// TIA Portal project "inzynierka2" (V17)

(* hardware
DEVICE "S7-1500/ET200MP station_1"  S7-1500 station
   slot 0: "Rail_0"  Rack  6ES7 590-1***0-0AA0
   slot 1: "PLC_1"  CPU 1513-1 PN  6ES7 513-1AL00-0AB0  V1.1
      slot 3: "CPU display_1"  6ES7591-1XA00-0AA0
      slot 32768: "PROFINET interface_1"  X1
DEVICE "GSD device_1"  GSD.Device.PN
   slot 0: "Rack"  Rack  V1.0
   slot 0: "CPX"  CPX-RC  TN 197330  V3.2.24
      slot 0: "CPX-RC"  CPX-RC
      slot 1: "PN-IO Interface"  PN-IO Interface
         slot 1: "Port 1"  Port 1
         slot 2: "Port 2"  Port 2
   slot 1: "FB34 PNIO Module (RC) [8IB/8OB]_1"  FB34 PNIO Module (RC) [8IB/8OB]  TN 548751, CPX-FB34
      slot 0: "FB34 PNIO Module (RC) [8IB/8OB]"  FB34 PNIO Module (RC) [8IB/8OB]
DEVICE "HMI_1"  KTP700 Basic PN
   slot 0: "HMI_1"  KTP700 Basic PN  6AV2 123-2GB03-0AX0  15.0.0.0
   slot 1: "HMI_RT_1"  KTP700 Basic PN  6AV2 123-2GB03-0AX0  15.0.0.0
   slot 5: "HMI_1.IE_CP_1"  PROFINET Interface  15.0.0.0
      slot 1: "PROFINET Interface_1"  PROFINET Interface
         slot 1: "Port_1"  Port
*)

// ===== PLC "PLC_1"  CPU 1513-1 PN =====

VAR_GLOBAL   // PLC tag table "Default tag table"
   "System_Byte" AT %MB1 : Byte;
   "FirstScan" AT %M1.0 : Bool;
   "DiagStatusUpdate" AT %M1.1 : Bool;
   "AlwaysTRUE" AT %M1.2 : Bool;
   "AlwaysFALSE" AT %M1.3 : Bool;
   "Clock_Byte" AT %MB0 : Byte;
   "Clock_10Hz" AT %M0.0 : Bool;
   "Clock_5Hz" AT %M0.1 : Bool;
   "Clock_2.5Hz" AT %M0.2 : Bool;
   "Clock_2Hz" AT %M0.3 : Bool;
   "Clock_1.25Hz" AT %M0.4 : Bool;
   "Clock_1Hz" AT %M0.5 : Bool;
   "Clock_0.625Hz" AT %M0.6 : Bool;
   "Clock_0.5Hz" AT %M0.7 : Bool;
   "Tag_1" AT %M10.1 : Bool;
   "testowy" AT %MB20 : Byte;
   "testowy_out" AT %MB22 : Byte;
   "testowy2" AT %MB21 : Byte;
   "testowy_out2" AT %MB23 : Byte;
   "Tag_2" AT %IW0 : Word;
   "IB_MANOMETER1_2" AT %IB0 : Byte;
   "IB_MANOMETER1_1" AT %IB1 : Byte;
   "valves_out_1" AT %MB100 : Byte;
   "QB0_BYTE_OUT" AT %QB0 : Byte;
   "valves_out_2" AT %MB101 : Byte;
   "QB1_BYTE_OUT" AT %QB1 : Byte;
   "QB2_BYTE_VALVE_OPEN_TO_SEND" AT %QB2 : Byte;
   "IB_MANOMETER3_2" AT %IB2 : Byte;
   "IB_MANOMETER3_1" AT %IB3 : Byte;
   "testint" AT %MW210 : Int;
   "testhmibool" AT %M212.0 : Bool;
   "IB_VALVE_STATE_1" AT %IB4 : Byte;
   "IB_VALVE_STATE_2" AT %IB5 : Byte;
   "IB_VALVE_STATE_3" AT %IB6 : Byte;
   "IB_VALVE_STATE_4" AT %IB7 : Byte;
   "Tag_3" AT %IB8 : Byte;
END_VAR

DATA_BLOCK "DB_send_rcv"   // DB1
{ S7_Optimized_Access := 'TRUE' }
VERSION : 0.1
   VAR
      przesuniecie : USInt;
      BAJT1 : Byte;
      BAJT2 : Byte;
      MANOMETER1_VALUE : Real;
      MANOMETER3_VALUE : Real;
      VALVE_OPEN_PERCENT : Int;
   END_VAR
BEGIN
END_DATA_BLOCK

DATA_BLOCK "DB_valves"   // DB2
{ S7_Optimized_Access := 'TRUE' }
VERSION : 0.1
   VAR
      VALVEMODE : Int := 1;
      TYPE_OF_2ND_INERTIA : Int := 1;
      VALVE_AUTO : Bool := TRUE;
      VALVE_MODE_STATE_ERR : Word;
      testbyte1 : Byte;
      testbyte2 : Byte;
      VALVE_STATE_CORRECT : Int;
      prop_display : Real;
   END_VAR
BEGIN
END_DATA_BLOCK

DATA_BLOCK "DB_PID"   // DB4
{ S7_Optimized_Access := 'TRUE' }
VERSION : 0.1
   VAR
      SETPOINT : Real;
      PID_OUT : Real;
      PID_COMPACT_AUTOTUNE : Bool := FALSE;
      PID_COMPACT_MANUAL_TUNE : Bool := TRUE;
      MANUAL_OUT : Real;
      PID_MANUALOUT : Bool := TRUE;
      PID_OUT_MAN : Real;
      MANUAL_LASTSTATE : Bool;
   END_VAR
BEGIN
END_DATA_BLOCK

FUNCTION "korekcja_bitow" : Void   // FC1, SCL
{ S7_Optimized_Access := 'TRUE' }
VERSION : 0.1
BEGIN
   "testowy_out" := ROR(IN := "testowy", N := "DB_send_rcv".przesuniecie);
END_FUNCTION

FUNCTION "rcv_pres" : Void   // FC2, SCL
{ S7_Optimized_Access := 'TRUE' }
VERSION : 0.1
   VAR_INPUT
      BYTE1 : Byte;
      BYTE2 : Byte;
   END_VAR
   VAR_OUTPUT
      OUT_PRES : Real;
   END_VAR
   VAR_TEMP
      TWOBYTES : Word;
      HI_PRES : Int;
   END_VAR
BEGIN
   #TWOBYTES:=(SHL(IN:=BYTE_TO_WORD(#BYTE1), N:=8) OR #BYTE2);
   #HI_PRES := WORD_TO_INT(#TWOBYTES);
   #OUT_PRES := INT_TO_REAL(#HI_PRES)/100.0;
END_FUNCTION

FUNCTION "valve_config" : Void   // FC3, SCL
{ S7_Optimized_Access := 'TRUE' }
VERSION : 0.1
   VAR_INPUT
      config : Int;   // 1:2nd inertia 2:extra container 3:all open 4:all close
      MODE_2ND : Int;   // TYPE OF 2ND INERTIA
      valve_autoconfig : Bool;
      valve_state1 : Byte;
      valve_state2 : Byte;
      valve_state3 : Byte;
      valve_state4 : Byte;
      valve_prop_sp : Real;
   END_VAR
   VAR_OUTPUT
      state_code : Word;   // 10:manual config 1X: config err
      valve_state_NB : Int;
      valve_prop_display : Real;
   END_VAR
   VAR_TEMP
      valve_config_nb : Int;
   END_VAR
   VAR CONSTANT
      config_ok : Bool;
   END_VAR
BEGIN
   #valve_config_nb := #config;
   #valve_prop_display := #valve_prop_sp / 25.0;



   IF NOT #valve_autoconfig THEN

       #valve_config_nb := 0;

   END_IF;


   CASE #valve_config_nb OF
       1:
           IF #MODE_2ND=1 THEN
               "valves_out_1" := 2#10001110; //2#10001110;
               "valves_out_2" := 2#11001011; // 2#11111000;

               IF #valve_state1=16#61 AND #valve_state2=16#1A AND #valve_state3=16#C3 AND #valve_state4=16#52 THEN
                   #state_code := 16#1;
                   #valve_state_NB := 1;
               ELSE
                   #state_code := 16#11;
                   #valve_state_NB := 2;
               END_IF
               ;
           ELSIF #MODE_2ND=2 THEN

               "valves_out_1" := 2#00110110; //2#10001110;
               "valves_out_2" := 2#11001101; // 2#11111000;

               IF #valve_state1 = 16#61 AND #valve_state2 = 16#29 AND #valve_state3 = 16#96 AND #valve_state4 = 16#34 THEN
                   #state_code := 16#1;
                   #valve_state_NB := 1;
               ELSE
                   #state_code := 16#11;
                   #valve_state_NB := 2;
               END_IF
               ;

           END_IF;




           ;

       2:

               "valves_out_1" := 2#00011110;
               "valves_out_2" := 2#11000101;
               IF #valve_state1=16#61 AND #valve_state2=16#38 AND #valve_state3=16#87 AND #valve_state4=16#25 THEN
                   #state_code := 16#2;
                   #valve_state_NB := 1;
               ELSE
                   #state_code := 16#12;
                   #valve_state_NB := 2;
               END_IF
               ;









       3:

           "valves_out_1" := 2#00000000;
           "valves_out_2" := 2#00000000;


           IF #valve_state1=16#07 AND #valve_state2=16#0B AND #valve_state3=16#0F AND #valve_state4=16#07 THEN
               #state_code := 16#3;
               #valve_state_NB := 1;
           ELSE
               #state_code := 16#13;
               #valve_state_NB := 2;
           END_IF
           ;

       4:
           "valves_out_1" := 2#11111111;

           "valves_out_2" := 2#11111111;

           IF #valve_state1=16#70 AND #valve_state2=16#38 AND #valve_state3=16#F0 AND #valve_state4=16#70 THEN
               #state_code := 16#4;
               #valve_state_NB := 1;
           ELSE
               #state_code := 16#14;
               #valve_state_NB := 2;
           END_IF
           ;


       ELSE

           #state_code := 16#10;
           #valve_state_NB := 3;
           ;
   END_CASE;
END_FUNCTION

FUNCTION "valves_set" : Void   // FC4, SCL
{ S7_Optimized_Access := 'TRUE' }
VERSION : 0.1
BEGIN

   "QB0_BYTE_OUT" := "valves_out_1";
   "QB1_BYTE_OUT" := "valves_out_2";
END_FUNCTION

FUNCTION "send_valve" : Void   // FC5, SCL
{ S7_Optimized_Access := 'TRUE' }
VERSION : 0.1
   VAR_INPUT
      DATA_TO_SEND : Real;
   END_VAR
   VAR_OUTPUT
      BYTE1 : Byte;
   END_VAR
   VAR_TEMP
      temp_byte : Byte;
      PRESS_CONVERT : Int;
      TEMP_DATA_TO_SEND : Real;
   END_VAR
BEGIN
   #TEMP_DATA_TO_SEND := #DATA_TO_SEND * 25.0;
   #PRESS_CONVERT := REAL_TO_INT(#TEMP_DATA_TO_SEND);
   #temp_byte := INT_TO_BYTE(#PRESS_CONVERT);
   #BYTE1 := #temp_byte;
END_FUNCTION

FUNCTION "mannual_out_valve" : Void   // FC6, SCL
{ S7_Optimized_Access := 'TRUE' }
VERSION : 0.1
   VAR_INPUT
      manual_value : Real;
   END_VAR
   VAR_OUTPUT
      manual_out_scal : Real;
   END_VAR
BEGIN
   #manual_out_scal := #manual_value * 25.0;
   //"DB_PID".SETPOINT := #manual_value;
END_FUNCTION

ORGANIZATION_BLOCK "Main"   // OB1, LAD, ProgramCycle
TITLE = "Main Program Sweep (Cycle)"
{ S7_Optimized_Access := 'TRUE' }
VERSION : 0.1
   VAR_INPUT
      Initial_Call : Bool;   // Initial call of this OB
      Remanence : Bool;   // =True, if remanent data are available
   END_VAR
   VAR_TEMP   // added for the SCL form of the ladder/FBD networks
      _w1 : Bool;
   END_VAR
BEGIN

REGION Network 1
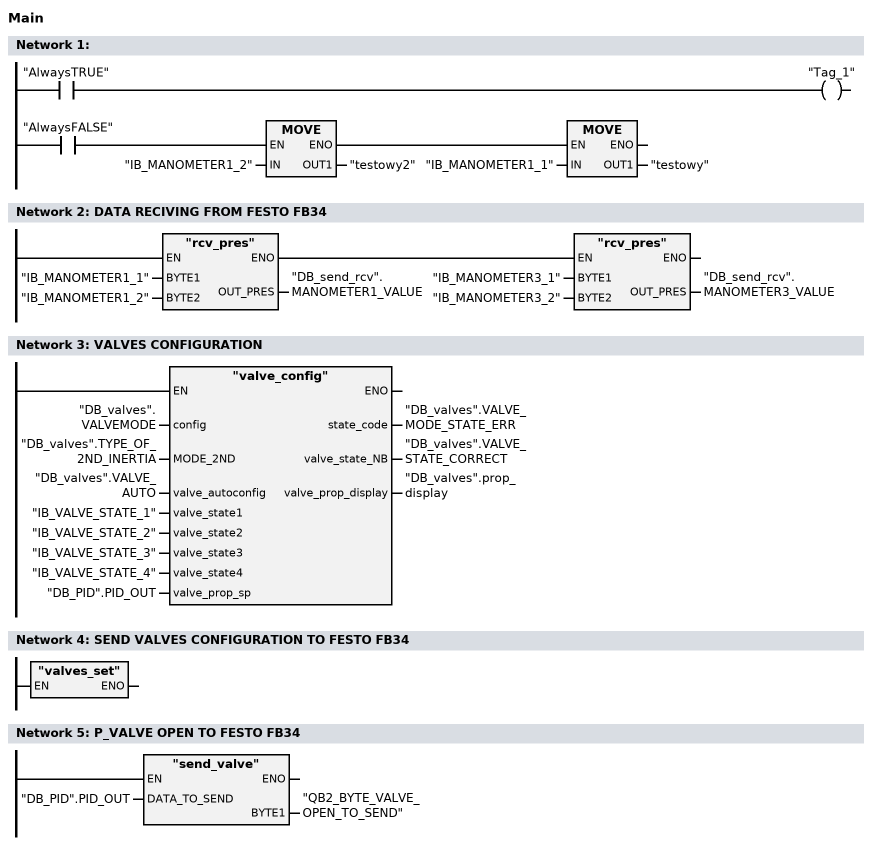
   RUNG wire#powerrail
      Contact( "AlwaysTRUE" )
      Coil( "Tag_1" )
   END_RUNG
   RUNG wire#powerrail
      Contact( "AlwaysFALSE" )
      Move(in := "IB_MANOMETER1_2", out1 => "testowy2")
      Move(in := "IB_MANOMETER1_1", out1 => "testowy")
   END_RUNG
   // the same network as SCL:
   "Tag_1" := "AlwaysTRUE";
   IF "AlwaysFALSE" THEN
       "testowy2" := "IB_MANOMETER1_2";
       "testowy" := "IB_MANOMETER1_1";
   END_IF;
END_REGION

REGION Network 2: DATA RECIVING FROM FESTO FB34
   RUNG wire#powerrail
      "rcv_pres"(BYTE1 := "IB_MANOMETER1_1", BYTE2 := "IB_MANOMETER1_2", OUT_PRES => "DB_send_rcv".MANOMETER1_VALUE)
      "rcv_pres"(BYTE1 := "IB_MANOMETER3_1", BYTE2 := "IB_MANOMETER3_2", OUT_PRES => "DB_send_rcv".MANOMETER3_VALUE)
   END_RUNG
   // the same network as SCL:
   "rcv_pres"(BYTE1 := "IB_MANOMETER1_1",
              BYTE2 := "IB_MANOMETER1_2",
              OUT_PRES => "DB_send_rcv".MANOMETER1_VALUE,
              ENO => #_w1);
   IF #_w1 THEN
       "rcv_pres"(BYTE1 := "IB_MANOMETER3_1",
                  BYTE2 := "IB_MANOMETER3_2",
                  OUT_PRES => "DB_send_rcv".MANOMETER3_VALUE);
   END_IF;
END_REGION

REGION Network 3: VALVES CONFIGURATION
   RUNG wire#powerrail
      "valve_config"(config := "DB_valves".VALVEMODE, MODE_2ND := "DB_valves".TYPE_OF_2ND_INERTIA, valve_autoconfig := "DB_valves".VALVE_AUTO, valve_state1 := "IB_VALVE_STATE_1", valve_state2 := "IB_VALVE_STATE_2", valve_state3 := "IB_VALVE_STATE_3", valve_state4 := "IB_VALVE_STATE_4", valve_prop_sp := "DB_PID".PID_OUT, state_code => "DB_valves".VALVE_MODE_STATE_ERR, valve_state_NB => "DB_valves".VALVE_STATE_CORRECT, valve_prop_display => "DB_valves".prop_display)
   END_RUNG
   // the same network as SCL:
   "valve_config"(config := "DB_valves".VALVEMODE,
                  MODE_2ND := "DB_valves".TYPE_OF_2ND_INERTIA,
                  valve_autoconfig := "DB_valves".VALVE_AUTO,
                  valve_state1 := "IB_VALVE_STATE_1",
                  valve_state2 := "IB_VALVE_STATE_2",
                  valve_state3 := "IB_VALVE_STATE_3",
                  valve_state4 := "IB_VALVE_STATE_4",
                  valve_prop_sp := "DB_PID".PID_OUT,
                  state_code => "DB_valves".VALVE_MODE_STATE_ERR,
                  valve_state_NB => "DB_valves".VALVE_STATE_CORRECT,
                  valve_prop_display => "DB_valves".prop_display);
END_REGION

REGION Network 4: SEND VALVES CONFIGURATION TO FESTO FB34
   RUNG wire#powerrail
      "valves_set"()
   END_RUNG
   // the same network as SCL:
   "valves_set"();
END_REGION

REGION Network 5: P_VALVE OPEN TO FESTO FB34
   RUNG wire#powerrail
      "send_valve"(DATA_TO_SEND := "DB_PID".PID_OUT, BYTE1 => "QB2_BYTE_VALVE_OPEN_TO_SEND")
   END_RUNG
   // the same network as SCL:
   "send_valve"(DATA_TO_SEND := "DB_PID".PID_OUT, BYTE1 => "QB2_BYTE_VALVE_OPEN_TO_SEND");
END_REGION
END_ORGANIZATION_BLOCK

ORGANIZATION_BLOCK "PID_block"   // OB30, LAD, CyclicInterrupt
{ S7_Optimized_Access := 'TRUE' }
VERSION : 0.1
   VAR_INPUT
      Initial_Call : Bool;   // Initial call of this OB
      Event_Count : Int;   // Events discarded
   END_VAR
   VAR_TEMP   // added for the SCL form of the ladder/FBD networks
      _w1 : Bool;
   END_VAR
BEGIN

REGION Network 1: bez udezeniowe
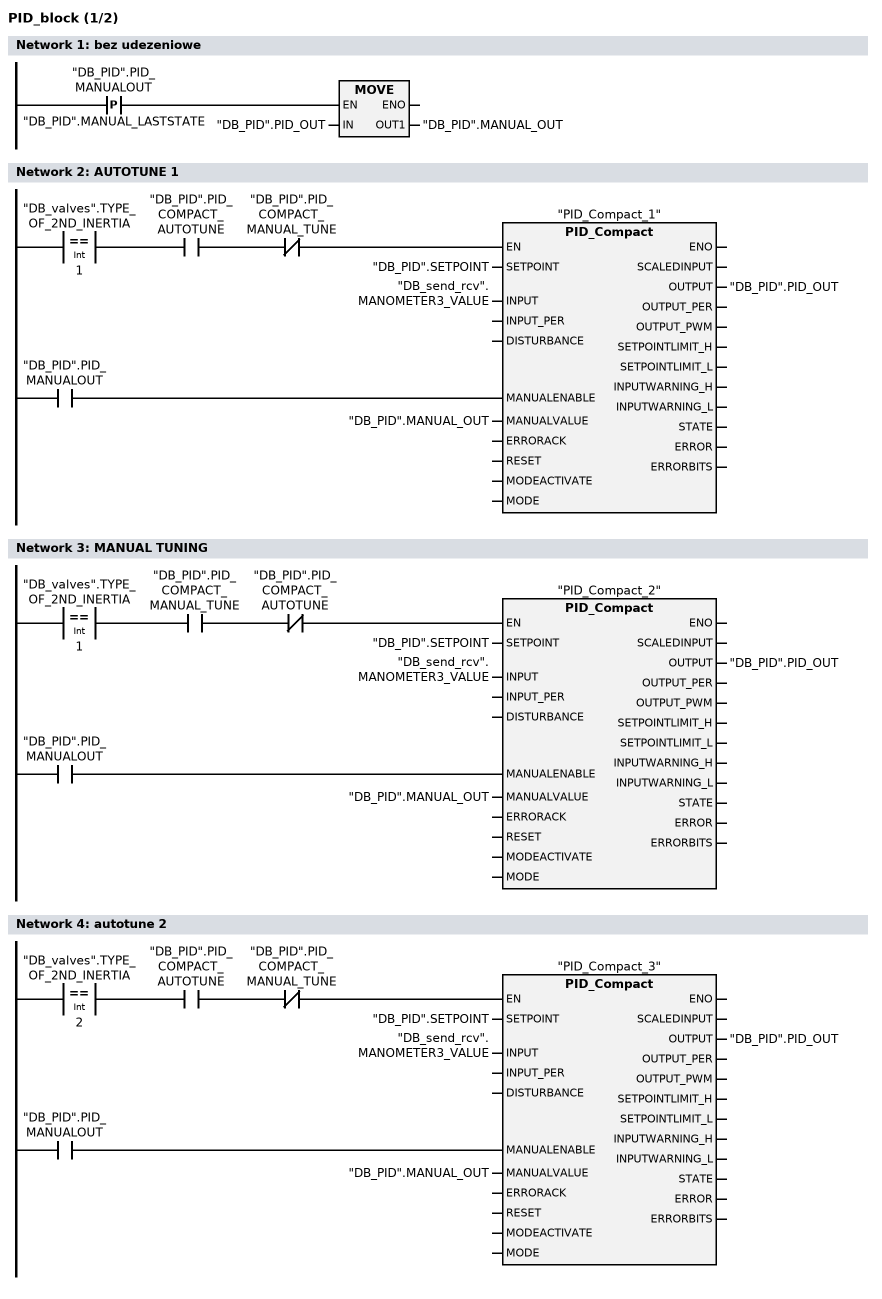
   RUNG wire#powerrail
      P_Contact(operand := "DB_PID".PID_MANUALOUT, bit := "DB_PID".MANUAL_LASTSTATE)
      Move(in := "DB_PID".PID_OUT, out1 => "DB_PID".MANUAL_OUT)
   END_RUNG
   // the same network as SCL:
   #_w1 := "DB_PID".PID_MANUALOUT AND NOT "DB_PID".MANUAL_LASTSTATE;   // rising edge of "DB_PID".PID_MANUALOUT
   "DB_PID".MANUAL_LASTSTATE := "DB_PID".PID_MANUALOUT;
   IF #_w1 THEN "DB_PID".MANUAL_OUT := "DB_PID".PID_OUT; END_IF;
END_REGION

REGION Network 2: AUTOTUNE 1
   IF ("DB_valves".TYPE_OF_2ND_INERTIA = 1) AND "DB_PID".PID_COMPACT_AUTOTUNE AND NOT "DB_PID".PID_COMPACT_MANUAL_TUNE THEN
       "PID_Compact_1"(Setpoint := "DB_PID".SETPOINT,   // PID_Compact
                       Input := "DB_send_rcv".MANOMETER3_VALUE,
                       ManualEnable := "DB_PID".PID_MANUALOUT,
                       ManualValue := "DB_PID".MANUAL_OUT,
                       Output => "DB_PID".PID_OUT);
   END_IF;
END_REGION

REGION Network 3: MANUAL TUNING
   IF ("DB_valves".TYPE_OF_2ND_INERTIA = 1) AND "DB_PID".PID_COMPACT_MANUAL_TUNE AND NOT "DB_PID".PID_COMPACT_AUTOTUNE THEN
       "PID_Compact_2"(Setpoint := "DB_PID".SETPOINT,   // PID_Compact
                       Input := "DB_send_rcv".MANOMETER3_VALUE,
                       ManualEnable := "DB_PID".PID_MANUALOUT,
                       ManualValue := "DB_PID".MANUAL_OUT,
                       Output => "DB_PID".PID_OUT);
   END_IF;
END_REGION

REGION Network 4: autotune 2
   IF ("DB_valves".TYPE_OF_2ND_INERTIA = 2) AND "DB_PID".PID_COMPACT_AUTOTUNE AND NOT "DB_PID".PID_COMPACT_MANUAL_TUNE THEN
       "PID_Compact_3"(Setpoint := "DB_PID".SETPOINT,   // PID_Compact
                       Input := "DB_send_rcv".MANOMETER3_VALUE,
                       ManualEnable := "DB_PID".PID_MANUALOUT,
                       ManualValue := "DB_PID".MANUAL_OUT,
                       Output => "DB_PID".PID_OUT);
   END_IF;
END_REGION

REGION Network 5
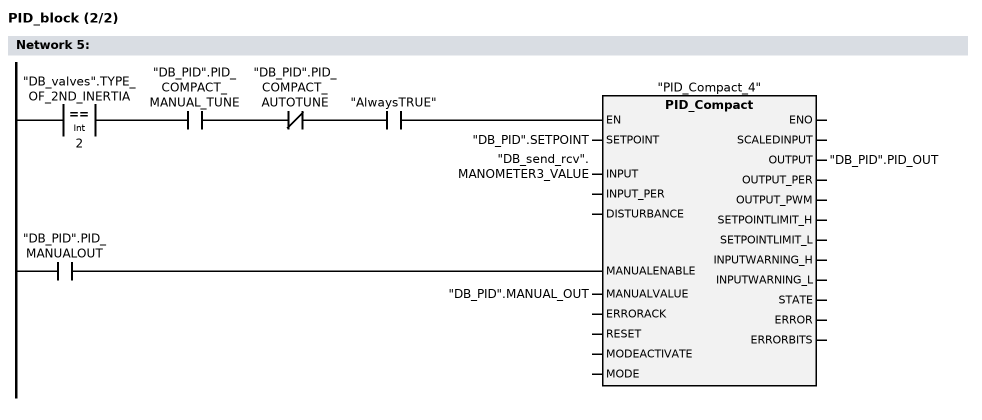
   IF ("DB_valves".TYPE_OF_2ND_INERTIA = 2) AND "DB_PID".PID_COMPACT_MANUAL_TUNE AND NOT "DB_PID".PID_COMPACT_AUTOTUNE AND "AlwaysTRUE" THEN
       "PID_Compact_4"(Setpoint := "DB_PID".SETPOINT,   // PID_Compact
                       Input := "DB_send_rcv".MANOMETER3_VALUE,
                       ManualEnable := "DB_PID".PID_MANUALOUT,
                       ManualValue := "DB_PID".MANUAL_OUT,
                       Output => "DB_PID".PID_OUT);
   END_IF;
END_REGION
END_ORGANIZATION_BLOCK

(* ===== HMI "HMI_RT_1" =====
system functions are stored by id; their names below are inferred from use
connection "HMI_Connection_1": ETHERNET, SMART_S7_1500_OMS

HMI tags "Default tag table"
   "Tag_ScreenNumber" : UInt, internal
   "testhmibool" : Bool = PLC testhmibool AT %M212.0, 1 s
   "DB_valves_VALVEMODE" : Int = PLC DB_valves.VALVEMODE, 1 s
   "DB_send_rcv_MANOMETER1_VALUE" : Real = PLC DB_send_rcv.MANOMETER1_VALUE, 1 s
   "DB_send_rcv_MANOMETER3_VALUE" : Real = PLC DB_send_rcv.MANOMETER3_VALUE, 1 s
   "DB_PID_SETPOINT" : Real = PLC DB_PID.SETPOINT, 1 s
   "DB_send_rcv_VALVE_OPEN_PERCENT" : Int = PLC DB_send_rcv.VALVE_OPEN_PERCENT, 1 s
   "DB_PID_PID_OUT" : Real = PLC DB_PID.PID_OUT, 1 s
   "DB_valves_VALVE_STATE_CORRECT" : Int = PLC DB_valves.VALVE_STATE_CORRECT, 1 s
   "DB_valves_VALVE_AUTO" : Bool = PLC DB_valves.VALVE_AUTO, 1 s
   "DB_PID_PID_COMPACT_AUTOTUNE" : Bool = PLC DB_PID.PID_COMPACT_AUTOTUNE, 1 s
   "DB_PID_PID_COMPACT_MANUAL_TUNE" : Bool = PLC DB_PID.PID_COMPACT_MANUAL_TUNE, 1 s
   "DB_PID_PID_MANUALOUT" : Bool = PLC DB_PID.PID_MANUALOUT, 1 s
   "DB_PID_MANUAL_OUT" : Real = PLC DB_PID.MANUAL_OUT, 1 s
   "DB_valves_prop_display" : Real = PLC DB_valves.prop_display, 1 s
   "DB_valves_TYPE_OF_2ND_INERTIA" : Int = PLC DB_valves.TYPE_OF_2ND_INERTIA, 1 s
   "PID_Compact_4_Retain_CtrlParams_Gain" : Real = PLC PID_Compact_4.Retain.CtrlParams.Gain, 1 s
   "PID_Compact_4_Retain_CtrlParams_Ti" : Real = PLC PID_Compact_4.Retain.CtrlParams.Ti, 1 s
   "PID_Compact_4_Retain_CtrlParams_Td" : Real = PLC PID_Compact_4.Retain.CtrlParams.Td, 1 s
   "PID_Compact_2_Retain_CtrlParams_Gain" : Real = PLC PID_Compact_2.Retain.CtrlParams.Gain, 1 s
   "PID_Compact_2_Retain_CtrlParams_Ti" : Real = PLC PID_Compact_2.Retain.CtrlParams.Ti, 1 s
   "PID_Compact_2_Retain_CtrlParams_Td" : Real = PLC PID_Compact_2.Retain.CtrlParams.Td, 1 s

text list "V_MODE": 1 '2ND INERTIA'; 2 '3RD INERTIA'; 3 'ALL OPEN'; 4 'ALL CLOSE'

text list "V_STATE": 1 'CORRECT'; 2 'ERROR'; 3 'MANUAL'

Template "Template_1" 800x480
   Button "Button_1" at 12,74 size 111x49; TextOff '2 rząd'
      on Press: SetTag("DB_valves_VALVEMODE", 1)
   Button "Button_2" at 12,74 size 120x49; TextOff '2ND INERTIA'
      on Press: SetTag("DB_valves_VALVEMODE", 1)
   Button "Button_3" at 12,127 size 120x49; TextOff '3RD INERTIA'
      on Press: SetTag("DB_valves_VALVEMODE", 2)
   IOField "Template_I/O field_1" at 12,210 size 120x42; FormatPattern 9.99
      ProcessValue <- "DB_send_rcv_MANOMETER1_VALUE"
   IOField "Template_I/O field_2" at 12,276 size 120x42; FormatPattern 9.99
      ProcessValue <- "DB_send_rcv_MANOMETER3_VALUE"
   IOField "Template_I/O field_3" at 12,343 size 120x43; FormatPattern 9.99
      ProcessValue <- "DB_PID_SETPOINT"
   SymbolicIOField "Template_Symbolic I/O field_1" at 564,3 size 176x39; TextOn '1'; TextOff '0'; TextList "V_MODE"
      ProcessValue <- "DB_valves_VALVEMODE"
   SymbolicIOField "Template_Symbolic I/O field_2" at 168,3 size 96x39; TextOn '1'; TextOff '0'; TextList "V_STATE"
      ProcessValue <- "DB_valves_VALVE_STATE_CORRECT"
   TextField "Template_Text field_1" at 466,11 size 59x23; Text 'MODE:'
   TextField "Template_Text field_2" at 54,11 size 74x23; Text 'VALVES:'
   TextField "Template_Text field_3" at 41,181 size 63x23; Text 'INPUT'
   TextField "Template_Text field_4" at 59,252 size 27x23; Text 'PV'
   TextField "Template_Text field_5" at 28,319 size 89x23; Text 'SETPOINT'
   Softkey "Softkey_F2" at 0,0 size 0x0
      on KeyDown: ActivateScreen("wykres", 0)
   Softkey "Softkey_F1" at 0,0 size 0x0
      on KeyDown: ActivateScreen("Root screen", 0)

screen "Root screen" 800x480, template "Template_2"
   on GenerateScreen: SetTag("Tag_ScreenNumber", 1)
   GraphicView "Graphic view_7" at 612,127 size 127x33; Picture "Graphic_2"
   GraphicView "Graphic view_6" at 191,123 size 127x33; Picture "Graphic_2"
   GraphicView "Graphic view_4" at 419,127 size 127x33; Picture "Graphic_2"
   GraphicView "Graphic view_1" at 290,43 size 158x195; Picture "Graphic_1"
   GraphicView "Graphic view_2" at 522,78 size 105x126; Picture "Graphic_1"
   GraphicView "Graphic view_3" at 679,106 size 62x70; Picture "Graphic_1"
   GraphicView "Graphic view_5" at 86,64 size 117x103; Picture "Graphic_3"
   IOField "Template_I/O field_1" at 118,174 size 54x38; FormatPattern 9.99
      ProcessValue <- "DB_send_rcv_MANOMETER1_VALUE"
   IOField "Template_I/O field_2" at 548,122 size 54x38; FormatPattern 9.99
      ProcessValue <- "DB_send_rcv_MANOMETER3_VALUE"
   IOField "Template_I/O field_3" at 548,239 size 54x38; FormatPattern 9.99
      ProcessValue <- "DB_PID_SETPOINT"
   GraphicView "Graphic view_12" at 379,234 size 48x48; Picture "Graphic_8"
   GraphicView "Graphic view_14" at 551,192 size 48x48; Picture "Graphic_10"
   GraphicView "Graphic view_8" at 507,234 size 48x48; Picture "Graphic_8"
   TextField "Text field_1" at 428,247 size 89x23; Text 'SETPOINT'
   GraphicView "Graphic view_9" at 8,124 size 83x80; Picture "Graphic_12"
   IOField "Template_I/O field_4" at 5,52 size 75x38; FormatPattern 9.99
      ProcessValue <- "DB_PID_PID_OUT"
   GraphicView "Graphic view_10" at 94,47 size 48x48; Picture "Graphic_8"
   Circle "Circle_1" at 25,282 size 28x28
      Appearance <- "DB_valves_VALVE_STATE_CORRECT"
   TextField "Text field_3" at 70,285 size 152x23; Text 'VALVES CORRECT'
   Button "Button_1" at 655,219 size 111x49; TextOff '2 rząd'
      on Press: SetTag("DB_valves_VALVEMODE", 1)
   Button "Button_2" at 650,219 size 120x49; TextOff '2ND INERTIA'
      on Press: SetTag("DB_valves_VALVEMODE", 1)
   Button "Button_3" at 650,280 size 120x49; TextOff '3RD INERTIA'
      on Press: SetTag("DB_valves_VALVEMODE", 2)
   Circle "Circle_2" at 358,54 size 23x23
      Visibility <- "DB_valves_VALVEMODE"
   Circle "Circle_3" at 563,86 size 23x23
      Visibility <- "DB_valves_VALVEMODE"
   Circle "Circle_4" at 699,111 size 23x23
      Visibility <- "DB_valves_VALVEMODE"
   Circle "Circle_5" at 358,54 size 23x23
      Visibility <- "DB_valves_TYPE_OF_2ND_INERTIA"
   Circle "Circle_7" at 563,86 size 23x23
      Visibility <- "DB_valves_TYPE_OF_2ND_INERTIA"
   Circle "Circle_8" at 563,86 size 23x23
      Visibility <- "DB_valves_TYPE_OF_2ND_INERTIA"
   Circle "Circle_9" at 699,111 size 23x23
      Visibility <- "DB_valves_TYPE_OF_2ND_INERTIA"

screen "wykres" 800x480, template "Template_1"
   TrendView "Trend view_1" at 172,44 size 603x383

screen "VALVES" 800x480, template "Template_2"
   Button "Button_2" at 331,116 size 139x49; TextOff '2ND INERTIA'
      on Press: SetTag("DB_valves_VALVEMODE", 1)
   Button "Button_3" at 331,193 size 139x49; TextOff '3RD INERTIA'
      on Press: SetTag("DB_valves_VALVEMODE", 2)
   Button "Button_5" at 331,270 size 139x49; TextOff 'ALL OPEN'
      on Press: SetTag("DB_valves_VALVEMODE", 3)
   Button "Button_6" at 331,348 size 139x49; TextOff 'ALL CLOSE'
      on Press: SetTag("DB_valves_VALVEMODE", 4)
   Switch "Switch_1" at 621,270 size 139x49; CaptionText 'Switch'; TextOff 'OFF'; TextOn 'ON'
      ProcessValue <- "DB_valves_VALVE_AUTO"
   TextField "Text field_1" at 598,234 size 188x28; Text 'VALVES SET AUTO'
   TextField "Text field_2" at 326,80 size 149x28; Text 'VALVES MODE'
   TextField "Text field_3" at 47,80 size 109x28; Text 'PID MODE'
   Button "Button_8" at 29,116 size 139x49; TextOff 'AUTO TUNE'
      on Press: SetBit("DB_PID_PID_COMPACT_AUTOTUNE"); ResetBit("DB_PID_PID_COMPACT_MANUAL_TUNE")
      Appearance <- "DB_PID_PID_COMPACT_AUTOTUNE"
   Button "Button_9" at 29,193 size 139x49; TextOff 'MANUAL TUNE'
      on Press: SetBit("DB_PID_PID_COMPACT_MANUAL_TUNE"); ResetBit("DB_PID_PID_COMPACT_AUTOTUNE")
      Appearance <- "DB_PID_PID_COMPACT_MANUAL_TUNE"
   Button "Button_1" at 29,270 size 139x49; TextOff 'MANUAL'
      Appearance <- "DB_PID_PID_MANUALOUT"
      on Press: InvertBit("DB_PID_PID_MANUALOUT")
   GraphicView "Graphic view_8" at 164,271 size 48x48; Picture "Graphic_8"
   IOField "I/O field_1" at 209,270 size 80x49; FormatPattern 9.99
      ProcessValue <- "DB_PID_MANUAL_OUT"
   Button "Button_4" at 621,116 size 64x49; TextOff '1'
      on Press: SetTag("DB_valves_TYPE_OF_2ND_INERTIA", 1)
   Button "Button_7" at 696,116 size 64x49; TextOff '2'
      on Press: SetTag("DB_valves_TYPE_OF_2ND_INERTIA", 2)
   TextField "Text field_4" at 587,80 size 208x28; Text '2ND INERTIA MODE'

Template "Template_2" 800x480
   SymbolicIOField "Template_Symbolic I/O field_1" at 564,3 size 176x39; TextOff '0'; TextOn '1'; TextList "V_MODE"
      ProcessValue <- "DB_valves_VALVEMODE"
   SymbolicIOField "Template_Symbolic I/O field_2" at 168,3 size 96x39; TextOff '0'; TextOn '1'; TextList "V_STATE"
      ProcessValue <- "DB_valves_VALVE_STATE_CORRECT"
   TextField "Template_Text field_1" at 466,11 size 59x23; Text 'MODE:'
   TextField "Template_Text field_2" at 54,11 size 74x23; Text 'VALVES:'

screen "PID" 800x480, template "Template_2"
   IOField "I/O field_1" at 583,150 size 96x32; FormatPattern s999999999.999
      ProcessValue <- "PID_Compact_4_Retain_CtrlParams_Gain"
   IOField "I/O field_2" at 584,226 size 96x32; FormatPattern s999999999.999
      ProcessValue <- "PID_Compact_4_Retain_CtrlParams_Ti"
   IOField "I/O field_3" at 587,302 size 96x32; FormatPattern s999999999.999
      ProcessValue <- "PID_Compact_4_Retain_CtrlParams_Td"
   IOField "I/O field_4" at 119,150 size 96x32; FormatPattern s999999999.999
      ProcessValue <- "PID_Compact_2_Retain_CtrlParams_Gain"
   IOField "I/O field_5" at 119,226 size 96x32; FormatPattern s999999999.999
      ProcessValue <- "PID_Compact_2_Retain_CtrlParams_Ti"
   IOField "I/O field_6" at 119,302 size 96x32; FormatPattern s999999999.999
      ProcessValue <- "PID_Compact_2_Retain_CtrlParams_Td"
   TextField "Text field_1" at 142,73 size 50x23; Text 'PID 1'
   TextField "Text field_2" at 606,73 size 50x23; Text 'PID 2'
   TextField "Text field_3" at 143,130 size 48x23; Text 'GAIN'
   TextField "Text field_4" at 157,206 size 21x23; Text 'Ti'
   TextField "Text field_5" at 154,282 size 26x23; Text 'Td'
   TextField "Text field_6" at 607,130 size 48x23; Text 'GAIN'
   TextField "Text field_7" at 621,206 size 21x23; Text 'Ti'
   TextField "Text field_8" at 618,282 size 26x23; Text 'Td'
*)